// TIA Portal project "Plc_KTKDL" (V19)

(* hardware
DEVICE "S7-1200 station_1"  S7-1200 Station
   slot 0: "Rack_0"  S7-1200 Rack  Rack  V1.0
   slot 1: "PLC_1"  CPU 1214C DC/DC/DC  6ES7 214-1AG40-0XB0  V4.0
DEVICE "PC-System_1"  SIMATIC PC station
   slot 0: "SIMATIC PC station"  Rail  SIMATIC PC-Station  V1.0
      slot 125: "Stationmanager"  Station_Manager  V6.0.4
   slot 1: "HMI_RT_1"  WinCC Unified PC RT  6AV2 155-xxxxx-xxxx  19.0.0.0
   slot 2: "IE general_1"  IE General  IE_CP  V8.2.0
      slot 1: "PROFINET interface"  IEGeneral.Interface.8.2.0
*)

// ===== PLC "PLC_1"  CPU 1214C DC/DC/DC =====

VAR_GLOBAL   // PLC tag table "Default tag table"
   "Step_Lift_Pulse" AT %Q0.0 : Bool;
   "Step_Lift_Direction" AT %Q0.1 : Bool;
   "Step_Reach_Pulse" AT %Q0.4 : Bool;
   "Step_Reach_Direction" AT %Q0.5 : Bool;
   "Axis_1_Direction" AT %Q0.3 : Bool;
   "Axis_1_Pulse" AT %Q0.2 : Bool;
   "Step_Lift_Homing switch" AT %I0.0 : Bool;
END_VAR

VAR_GLOBAL   // PLC tag table "Input"
   "SensorHome" AT %M0.1 : Bool;
END_VAR

TYPE "UDT"
   STRUCT
      Monitor : Struct
         Velocity : Real;
         Position : Real;
      END_STRUCT;
      Job : Struct
         Velocity : Real;
         Forwork : Bool;
         Backwork : Bool;
         Erorr : Bool;
      END_STRUCT;
      StaticAxis : Int;
   END_STRUCT;
END_TYPE

DATA_BLOCK "DB_Vị_trí_xe"   // DB2
{ S7_Optimized_Access := 'FALSE' }
VERSION : 0.1
   VAR
      "vị trí 1" : Bool;
      "vị trí 2" : Bool;
      "vị trí 3" : Bool;
      "vị trí 4" : Bool;
      "vị trí 5" : Bool;
      "vị trí 6" : Bool;
      "vị trí 7" : Bool;
      "vị trí 8" : Bool;
      tầng_1 : Bool;
      tầng_2 : Bool;
   END_VAR
BEGIN
END_DATA_BLOCK

DATA_BLOCK "P_Trig"   // DB3
{ S7_Optimized_Access := 'TRUE' }
VERSION : 0.1
   VAR
      CLK : Array[0..100] of Bool;
   END_VAR
BEGIN
END_DATA_BLOCK

DATA_BLOCK "DB_AxisPanel"   // DB5
{ S7_Optimized_Access := 'TRUE' }
VERSION : 0.1
   VAR
      Lift : "UDT";
      Rotation : "UDT";
      Reach : "UDT";
   END_VAR
BEGIN
END_DATA_BLOCK

DATA_BLOCK "DB_Operater"   // DB6
{ S7_Optimized_Access := 'FALSE' }
VERSION : 0.1
   VAR
      Confirm_Gửi : Bool;
      Confirm_Lấy : Bool;
      ConfirmRFID : Bool;
      Scada_Gửi_Xe : Bool;
      Scada_Lấy_Xe : Bool;
      Scada_RFID : Bool;
      Scada_Home_Lift : Bool;
      BackHome : Bool;
      "Auto/Man" : Bool;
      Static_Mode : Int;
   END_VAR
BEGIN
END_DATA_BLOCK

DATA_BLOCK "DB_Convert"   // DB14
{ S7_Optimized_Access := 'FALSE' }
VERSION : 0.1
   VAR
      Python : Struct
         Floor : Int := 0;
         Location : Int;
         Passcodeplc : Int;
         UID : Array[1..12] of String[14];
         Receive : String[14];
      END_STRUCT;
      Floor_Dic1 : Int;
      Floor_Dic2 : Int;
      Location : Int;
      Down : Int;
      Up : Int;
      Started : Bool;
   END_VAR
BEGIN
END_DATA_BLOCK

// folder: Step

DATA_BLOCK "DB_Step"   // DB15
{ S7_Optimized_Access := 'TRUE' }
VERSION : 0.1
   VAR
      Power : Bool;
      Home : Struct
         Lift : Bool;
         Rotation : Bool;
         Reach : Bool;
      END_STRUCT;
      HomeAll : Bool;
      ErorrHomeCode : Struct
         Lift : Word;
         Rotation : Word;
         Reach : Word;
      END_STRUCT;
      ErrorHome : Struct
         Lift : Bool;
         Rotation : Bool;
         Reach : Bool;
      END_STRUCT;
      ErorrAbsoluteCode : Struct
         Rotation : Word;
         Lift : Word;
         Reach : Word;
      END_STRUCT;
      ErrorAbsolute : Struct
         Lift : Bool;
         Rotation : Bool;
         Reach : Bool;
      END_STRUCT;
      ErrorJog : Struct
         Lift : Word;
         Rotation : Word;
         Reach : Word;
      END_STRUCT;
      Reset : Bool;
      PowerStarted : Bool;
      HomeStarted : Bool;
      DoneHome : Bool;
   END_VAR
BEGIN
END_DATA_BLOCK

DATA_BLOCK "DB_Scrips"   // DB45
{ S7_Optimized_Access := 'FALSE' }
VERSION : 0.1
   VAR
      Dic : Int;
      "Step" : Int;
      Velocity : Struct
         Lift : Int;
         Rotation : Int;
         Reach : Int;
      END_STRUCT;
      Position : Struct
         Lift : Int;
         Rotation : Int;
         Reach : Int;
      END_STRUCT;
      Excute : Struct
         Lift : Bool;
         Rotation : Bool;
         Reach : Bool;
      END_STRUCT;
      ExcuteReady : Bool;
      Cònirm2 : Bool;
      Cònirm1 : Bool;
      Busy : Bool;
   END_VAR
BEGIN
END_DATA_BLOCK

// folder: System blocks/Program resources

DATA_BLOCK "DelayStep3"   // DB11
{ S7_Optimized_Access := 'TRUE' }
AUTHOR : Simatic
FAMILY : IEC
NAME : IEC_TMR
VERSION : 1.0
// stored: InstanceOfName IEC_TIMER
"IEC_TIMER"
BEGIN
END_DATA_BLOCK

DATA_BLOCK "Delay2s"   // DB23
{ S7_Optimized_Access := 'TRUE' }
AUTHOR : Simatic
FAMILY : IEC
NAME : IEC_TMR
VERSION : 1.0
// stored: InstanceOfName IEC_TIMER
"IEC_TIMER"
BEGIN
END_DATA_BLOCK

DATA_BLOCK "DelayStep4"   // DB47
{ S7_Optimized_Access := 'TRUE' }
AUTHOR : Simatic
FAMILY : IEC
NAME : IEC_TMR
VERSION : 1.0
// stored: InstanceOfName IEC_TIMER
"IEC_TIMER"
BEGIN
END_DATA_BLOCK

DATA_BLOCK "Delay1s5"   // DB49
{ S7_Optimized_Access := 'TRUE' }
AUTHOR : Simatic
FAMILY : IEC
NAME : IEC_TMR
VERSION : 1.0
// stored: InstanceOfName IEC_TIMER
"IEC_TIMER"
BEGIN
END_DATA_BLOCK

DATA_BLOCK "DelayyStep3"   // DB50
{ S7_Optimized_Access := 'TRUE' }
AUTHOR : Simatic
FAMILY : IEC
NAME : IEC_TMR
VERSION : 1.0
// stored: InstanceOfName IEC_TIMER
"IEC_TIMER"
BEGIN
END_DATA_BLOCK

// folder: đầy , các logic tìm

DATA_BLOCK "DB_Tìm&&Xácnhan"   // DB1
{ S7_Optimized_Access := 'TRUE' }
VERSION : 0.1
   VAR
      Call_tìm_vị_trí : Bool;
      Call_tìm_tầng : Bool;
      Xác_nhận_vị_trí : DInt;
      Xác_nhận_tầng : DInt;
   END_VAR
BEGIN
END_DATA_BLOCK

DATA_BLOCK "DB_đầy"   // DB4
{ S7_Optimized_Access := 'TRUE' }
VERSION : 0.1
   VAR
      Tầng1 : Bool;
      Tầng2 : Bool;
   END_VAR
BEGIN
END_DATA_BLOCK

// folder: (top level)

DATA_BLOCK "Step_Lift"   // DB10, Motion_DB
{ S7_Optimized_Access := 'TRUE' }
AUTHOR : SIMATIC
FAMILY : BasicMC
NAME : TO_PosAx
VERSION : 4.0
// stored: InstanceOfName TO_PositioningAxis
"TO_PositioningAxis"
BEGIN
   // Axis.DirectionOutputEnabledCU = TRUE
   // Axis.OnlinePtoModeCU = 16#0000_0002
   // Axis.SelectedChannel2EnumCU = %Q0.1
   // Axis.SelectedChannel1EnumCU = %Q0.0
   // Pulse.MinDeltaDeltaFrequencyCU = 0.004
   // Pulse.MaxDeltaDeltaFrequencyCU = 1.0E+10
   // Pulse.MinDeltaFrequencyCU = 0.005
   // Pulse.MaxDeltaFrequencyCU = 9.5E+9
   // Pulse.MinFrequencyCU = 1.0
   // Pulse.MaxFrequencyCU = 100000.0
   // Pulse.OutputSourceCU = 16#0000_0000
   // Axis.SelectPTO = 0
   // Axis.LengthUnitNormalized.Distance = 1013
END_DATA_BLOCK

DATA_BLOCK "Step_Reach"   // DB12, Motion_DB
{ S7_Optimized_Access := 'TRUE' }
AUTHOR : SIMATIC
FAMILY : BasicMC
NAME : TO_PosAx
VERSION : 4.0
// stored: InstanceOfName TO_PositioningAxis
"TO_PositioningAxis"
BEGIN
   // Axis.DirectionOutputEnabledCU = TRUE
   // Axis.OnlinePtoModeCU = 16#0000_0002
   // Axis.SelectedChannel2EnumCU = %Q0.5
   // Axis.SelectedChannel1EnumCU = %Q0.4
   // Pulse.MinDeltaDeltaFrequencyCU = 0.004
   // Pulse.MaxDeltaDeltaFrequencyCU = 1.0E+10
   // Pulse.MinDeltaFrequencyCU = 0.005
   // Pulse.MaxDeltaFrequencyCU = 9.5E+9
   // Pulse.MinFrequencyCU = 1.0
   // Pulse.MaxFrequencyCU = 30000.0
   // Pulse.OutputSourceCU = 16#0000_0000
   // Axis.SelectPTO = 1
   // Axis.OnlinePtoIndexCU = 1
   // Axis.LengthUnitNormalized.Distance = 1013
END_DATA_BLOCK

DATA_BLOCK "Step_Rotation"   // DB13, Motion_DB
{ S7_Optimized_Access := 'TRUE' }
AUTHOR : SIMATIC
FAMILY : BasicMC
NAME : TO_PosAx
VERSION : 4.0
// stored: InstanceOfName TO_PositioningAxis
"TO_PositioningAxis"
BEGIN
   // Axis.LengthUnitNormalized.Distance = 1005
   // Axis.LengthUnit.LastDistance = 1005
   // Axis.DirectionOutputEnabledCU = TRUE
   // Axis.OnlinePtoModeCU = 16#0000_0002
   // Axis.SelectedChannel2EnumCU = %Q0.3
   // Axis.SelectedChannel1EnumCU = %Q0.2
   // Pulse.MinDeltaDeltaFrequencyCU = 0.004
   // Pulse.MaxDeltaDeltaFrequencyCU = 1.0E+10
   // Pulse.MinDeltaFrequencyCU = 0.005
   // Pulse.MaxDeltaFrequencyCU = 9.5E+9
   // Pulse.MinFrequencyCU = 1.0
   // Pulse.MaxFrequencyCU = 100000.0
   // Pulse.OutputSourceCU = 16#0000_0000
   // Axis.SelectPTO = 2
   // Axis.OnlinePtoIndexCU = 2
END_DATA_BLOCK

FUNCTION "FC_SendPython" : Void   // FC1, LAD
{ S7_Optimized_Access := 'TRUE' }
VERSION : 0.1
BEGIN

REGION Network 1
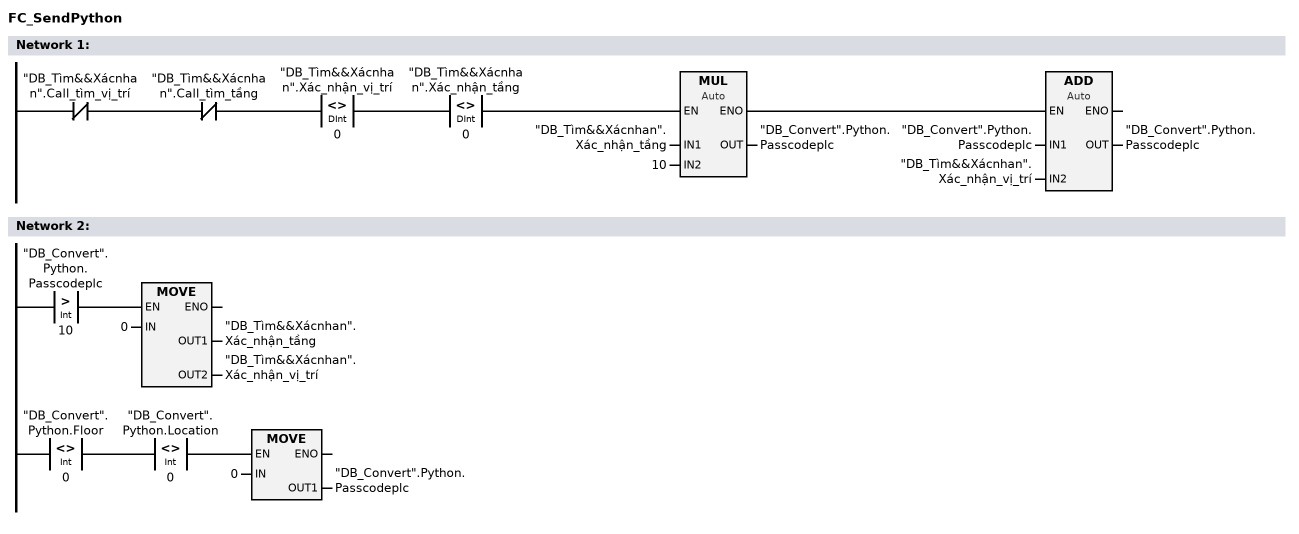
   RUNG wire#powerrail
      I_Contact( "DB_Tìm&&Xácnhan".Call_tìm_vị_trí )
      I_Contact( "DB_Tìm&&Xácnhan".Call_tìm_tầng )
      { S7_Templates := "SrcType := DInt" } NE_Contact(in1 := "DB_Tìm&&Xácnhan".Xác_nhận_vị_trí, in2 := 0)
      { S7_Templates := "SrcType := DInt" } NE_Contact(in1 := "DB_Tìm&&Xácnhan".Xác_nhận_tầng, in2 := 0)
      Mul(in1 := "DB_Tìm&&Xácnhan".Xác_nhận_tầng, in2 := 10, out => "DB_Convert".Python.Passcodeplc)
      Add(in1 := "DB_Convert".Python.Passcodeplc, in2 := "DB_Tìm&&Xácnhan".Xác_nhận_vị_trí, out => "DB_Convert".Python.Passcodeplc)
   END_RUNG
   // the same network as SCL:
   IF NOT "DB_Tìm&&Xácnhan".Call_tìm_vị_trí AND NOT "DB_Tìm&&Xácnhan".Call_tìm_tầng AND ("DB_Tìm&&Xácnhan".Xác_nhận_vị_trí <> 0) AND ("DB_Tìm&&Xácnhan".Xác_nhận_tầng <> 0) THEN
       "DB_Convert".Python.Passcodeplc := "DB_Tìm&&Xácnhan".Xác_nhận_tầng * 10;
       "DB_Convert".Python.Passcodeplc := "DB_Convert".Python.Passcodeplc + "DB_Tìm&&Xácnhan".Xác_nhận_vị_trí;
   END_IF;
END_REGION

REGION Network 2
   RUNG wire#powerrail
      { S7_Templates := "SrcType := Int" } GT_Contact(in1 := "DB_Convert".Python.Passcodeplc, in2 := 10)
      Move(in := 0, out1 => "DB_Tìm&&Xácnhan".Xác_nhận_tầng, out2 => "DB_Tìm&&Xácnhan".Xác_nhận_vị_trí)
   END_RUNG
   RUNG wire#powerrail
      { S7_Templates := "SrcType := Int" } NE_Contact(in1 := "DB_Convert".Python.Floor, in2 := 0)
      { S7_Templates := "SrcType := Int" } NE_Contact(in1 := "DB_Convert".Python.Location, in2 := 0)
      Move(in := 0, out1 => "DB_Convert".Python.Passcodeplc)
   END_RUNG
   // the same network as SCL:
   IF "DB_Convert".Python.Passcodeplc > 10 THEN
       "DB_Tìm&&Xácnhan".Xác_nhận_tầng := 0;
       "DB_Tìm&&Xácnhan".Xác_nhận_vị_trí := 0;
   END_IF;
   IF ("DB_Convert".Python.Floor <> 0) AND ("DB_Convert".Python.Location <> 0) THEN
       "DB_Convert".Python.Passcodeplc := 0;
   END_IF;
END_REGION
END_FUNCTION

FUNCTION "FC_Operater" : Void   // FC5, LAD
{ S7_Optimized_Access := 'TRUE' }
VERSION : 0.1
   VAR_TEMP   // added for the SCL form of the ladder/FBD networks
      _w1 : Bool;
      _w2 : Bool;
   END_VAR
BEGIN

REGION Network 1
   // chờ khi người dùng bấm rồi mới chạy
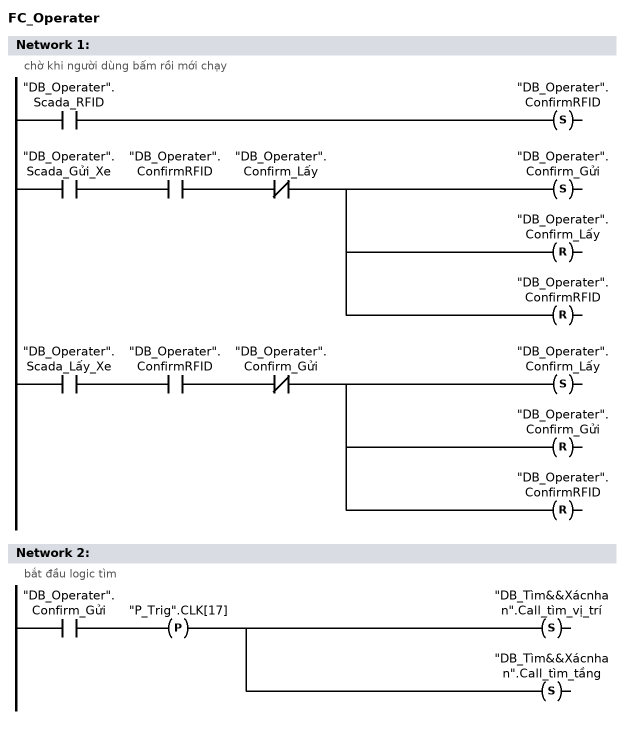
   RUNG wire#powerrail
      Contact( "DB_Operater".Scada_RFID )
      S_Coil( "DB_Operater".ConfirmRFID )
   END_RUNG
   RUNG wire#powerrail
      Contact( "DB_Operater".Scada_Gửi_Xe )
      Contact( "DB_Operater".ConfirmRFID )
      I_Contact( "DB_Operater".Confirm_Lấy )
      wire#w1
      S_Coil( "DB_Operater".Confirm_Gửi )
   END_RUNG
   RUNG wire#w1
      R_Coil( "DB_Operater".Confirm_Lấy )
   END_RUNG
   RUNG wire#w1
      R_Coil( "DB_Operater".ConfirmRFID )
   END_RUNG
   RUNG wire#powerrail
      Contact( "DB_Operater".Scada_Lấy_Xe )
      Contact( "DB_Operater".ConfirmRFID )
      I_Contact( "DB_Operater".Confirm_Gửi )
      wire#w2
      S_Coil( "DB_Operater".Confirm_Lấy )
   END_RUNG
   RUNG wire#w2
      R_Coil( "DB_Operater".Confirm_Gửi )
   END_RUNG
   RUNG wire#w2
      R_Coil( "DB_Operater".ConfirmRFID )
   END_RUNG
   // the same network as SCL:
   IF "DB_Operater".Scada_RFID THEN "DB_Operater".ConfirmRFID := TRUE; END_IF;
   IF "DB_Operater".Scada_Gửi_Xe AND "DB_Operater".ConfirmRFID AND NOT "DB_Operater".Confirm_Lấy THEN
       "DB_Operater".Confirm_Gửi := TRUE;
   END_IF;
   #_w1 := "DB_Operater".Scada_Gửi_Xe AND "DB_Operater".ConfirmRFID AND NOT "DB_Operater".Confirm_Lấy;
   IF #_w1 THEN
       "DB_Operater".Confirm_Lấy := FALSE;
       "DB_Operater".ConfirmRFID := FALSE;
   END_IF;
   IF "DB_Operater".Scada_Lấy_Xe AND "DB_Operater".ConfirmRFID AND NOT "DB_Operater".Confirm_Gửi THEN
       "DB_Operater".Confirm_Lấy := TRUE;
   END_IF;
   #_w2 := "DB_Operater".Scada_Lấy_Xe AND "DB_Operater".ConfirmRFID AND NOT "DB_Operater".Confirm_Gửi;
   IF #_w2 THEN
       "DB_Operater".Confirm_Gửi := FALSE;
       "DB_Operater".ConfirmRFID := FALSE;
   END_IF;
END_REGION

REGION Network 2
   // bắt đầu logic tìm
   RUNG wire#powerrail
      Contact( "DB_Operater".Confirm_Gửi )
      P_Trig( "P_Trig".CLK[17] )
      wire#w1
      S_Coil( "DB_Tìm&&Xácnhan".Call_tìm_vị_trí )
   END_RUNG
   RUNG wire#w1
      S_Coil( "DB_Tìm&&Xácnhan".Call_tìm_tầng )
   END_RUNG
   // the same network as SCL:
   #_w1 := "DB_Operater".Confirm_Gửi AND NOT "P_Trig".CLK[17];   // rising edge
   "P_Trig".CLK[17] := "DB_Operater".Confirm_Gửi;
   IF #_w1 THEN
       "DB_Tìm&&Xácnhan".Call_tìm_vị_trí := TRUE;
       "DB_Tìm&&Xácnhan".Call_tìm_tầng := TRUE;
   END_IF;
END_REGION
END_FUNCTION

FUNCTION "Fc_Convert" : Void   // FC7, LAD
{ S7_Optimized_Access := 'TRUE' }
VERSION : 0.1
BEGIN

REGION Network 1
   // chuyen quang duong di cua truc nang
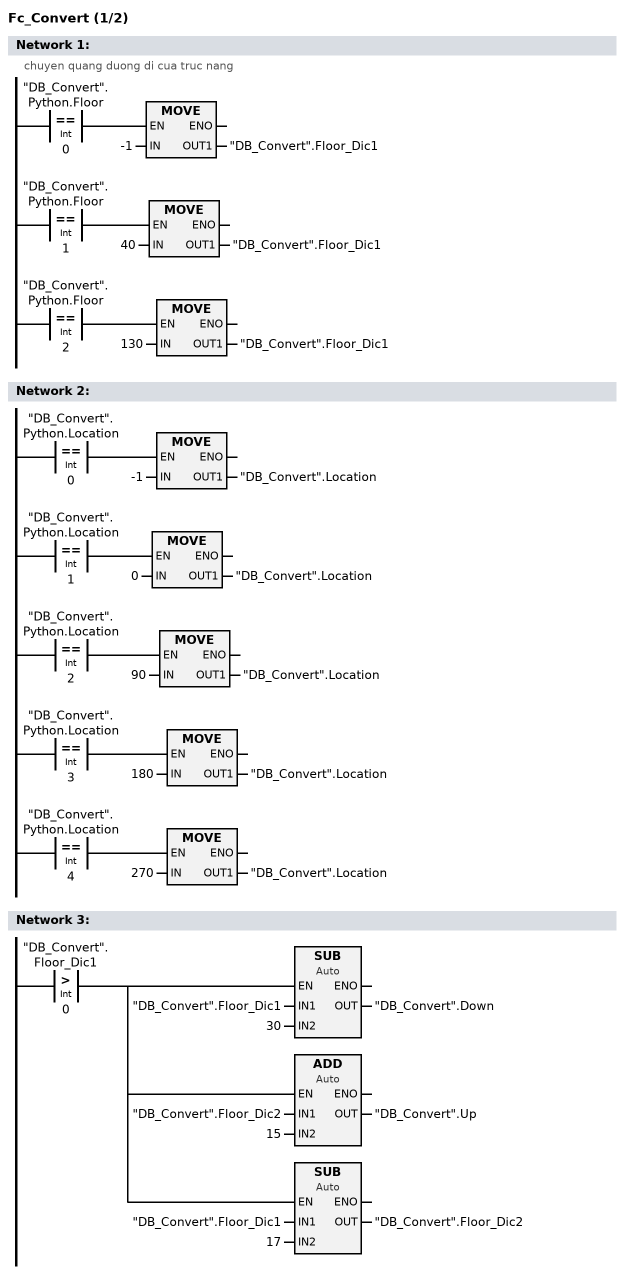
   RUNG wire#powerrail
      { S7_Templates := "SrcType := Int" } EQ_Contact(in1 := "DB_Convert".Python.Floor, in2 := 0)
      Move(in := -1, out1 => "DB_Convert".Floor_Dic1)
   END_RUNG
   RUNG wire#powerrail
      { S7_Templates := "SrcType := Int" } EQ_Contact(in1 := "DB_Convert".Python.Floor, in2 := 1)
      Move(in := 40, out1 => "DB_Convert".Floor_Dic1)
   END_RUNG
   RUNG wire#powerrail
      { S7_Templates := "SrcType := Int" } EQ_Contact(in1 := "DB_Convert".Python.Floor, in2 := 2)
      Move(in := 130, out1 => "DB_Convert".Floor_Dic1)
   END_RUNG
   // the same network as SCL:
   IF "DB_Convert".Python.Floor = 0 THEN "DB_Convert".Floor_Dic1 := -1; END_IF;
   IF "DB_Convert".Python.Floor = 1 THEN "DB_Convert".Floor_Dic1 := 40; END_IF;
   IF "DB_Convert".Python.Floor = 2 THEN "DB_Convert".Floor_Dic1 := 130; END_IF;
END_REGION

REGION Network 2
   RUNG wire#powerrail
      { S7_Templates := "SrcType := Int" } EQ_Contact(in1 := "DB_Convert".Python.Location, in2 := 0)
      Move(in := -1, out1 => "DB_Convert".Location)
   END_RUNG
   RUNG wire#powerrail
      { S7_Templates := "SrcType := Int" } EQ_Contact(in1 := "DB_Convert".Python.Location, in2 := 1)
      Move(in := 0, out1 => "DB_Convert".Location)
   END_RUNG
   RUNG wire#powerrail
      { S7_Templates := "SrcType := Int" } EQ_Contact(in1 := "DB_Convert".Python.Location, in2 := 2)
      Move(in := 90, out1 => "DB_Convert".Location)
   END_RUNG
   RUNG wire#powerrail
      { S7_Templates := "SrcType := Int" } EQ_Contact(in1 := "DB_Convert".Python.Location, in2 := 3)
      Move(in := 180, out1 => "DB_Convert".Location)
   END_RUNG
   RUNG wire#powerrail
      { S7_Templates := "SrcType := Int" } EQ_Contact(in1 := "DB_Convert".Python.Location, in2 := 4)
      Move(in := 270, out1 => "DB_Convert".Location)
   END_RUNG
   // the same network as SCL:
   IF "DB_Convert".Python.Location = 0 THEN "DB_Convert".Location := -1; END_IF;
   IF "DB_Convert".Python.Location = 1 THEN "DB_Convert".Location := 0; END_IF;
   IF "DB_Convert".Python.Location = 2 THEN "DB_Convert".Location := 90; END_IF;
   IF "DB_Convert".Python.Location = 3 THEN "DB_Convert".Location := 180; END_IF;
   IF "DB_Convert".Python.Location = 4 THEN "DB_Convert".Location := 270; END_IF;
END_REGION

REGION Network 3
   RUNG wire#powerrail
      { S7_Templates := "SrcType := Int" } GT_Contact(in1 := "DB_Convert".Floor_Dic1, in2 := 0)
      wire#w1
      Sub(in1 := "DB_Convert".Floor_Dic1, in2 := 30, out => "DB_Convert".Down)
   END_RUNG
   RUNG wire#w1
      Add(in1 := "DB_Convert".Floor_Dic2, in2 := 15, out => "DB_Convert".Up)
   END_RUNG
   RUNG wire#w1
      Sub(in1 := "DB_Convert".Floor_Dic1, in2 := 17, out => "DB_Convert".Floor_Dic2)
   END_RUNG
   // the same network as SCL:
   IF "DB_Convert".Floor_Dic1 > 0 THEN
       "DB_Convert".Down := "DB_Convert".Floor_Dic1 - 30;
       "DB_Convert".Up := "DB_Convert".Floor_Dic2 + 15;
       "DB_Convert".Floor_Dic2 := "DB_Convert".Floor_Dic1 - 17;
   END_IF;
END_REGION

REGION Network 4
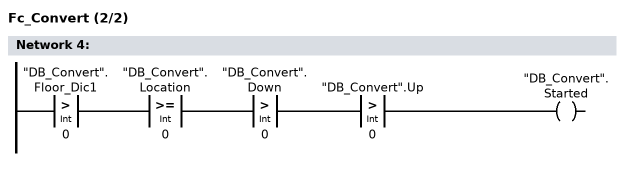
   RUNG wire#powerrail
      { S7_Templates := "SrcType := Int" } GT_Contact(in1 := "DB_Convert".Floor_Dic1, in2 := 0)
      { S7_Templates := "SrcType := Int" } GE_Contact(in1 := "DB_Convert".Location, in2 := 0)
      { S7_Templates := "SrcType := Int" } GT_Contact(in1 := "DB_Convert".Down, in2 := 0)
      { S7_Templates := "SrcType := Int" } GT_Contact(in1 := "DB_Convert".Up, in2 := 0)
      Coil( "DB_Convert".Started )
   END_RUNG
   // the same network as SCL:
   "DB_Convert".Started := ("DB_Convert".Floor_Dic1 > 0) AND ("DB_Convert".Location >= 0) AND ("DB_Convert".Down > 0) AND ("DB_Convert".Up > 0);
END_REGION
END_FUNCTION

FUNCTION "FC_Manual" : Void   // FC9, LAD
{ S7_Optimized_Access := 'TRUE' }
VERSION : 0.1
   VAR_TEMP   // added for the SCL form of the ladder/FBD networks
      _w1 : Bool;
   END_VAR
BEGIN

REGION Network 1
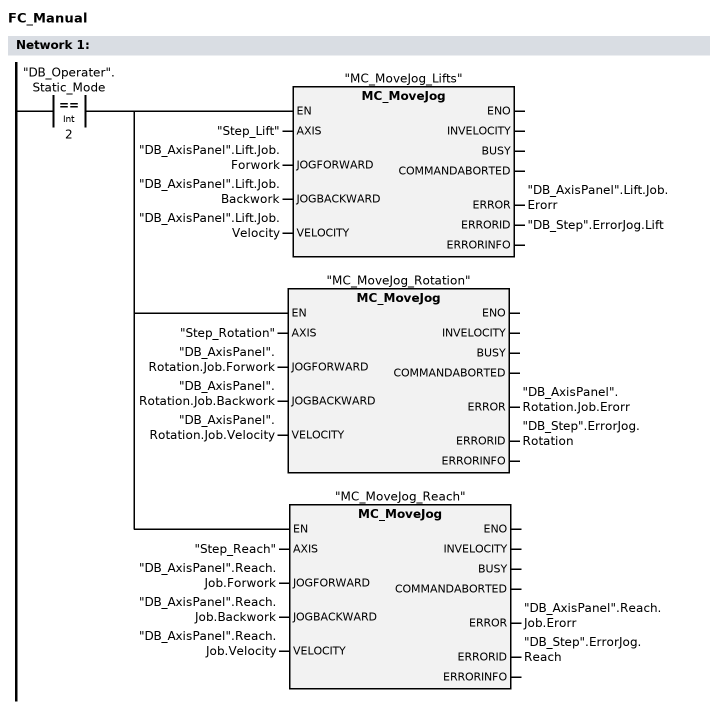
   #_w1 := "DB_Operater".Static_Mode = 2;
   IF #_w1 THEN
       "MC_MoveJog_Lifts"(Axis := "Step_Lift",   // MC_MoveJog
                          JogForward := "DB_AxisPanel".Lift.Job.Forwork,
                          JogBackward := "DB_AxisPanel".Lift.Job.Backwork,
                          Velocity := "DB_AxisPanel".Lift.Job.Velocity,
                          Error => "DB_AxisPanel".Lift.Job.Erorr,
                          ErrorID => "DB_Step".ErrorJog.Lift);
       "MC_MoveJog_Rotation"(Axis := "Step_Rotation",   // MC_MoveJog
                             JogForward := "DB_AxisPanel".Rotation.Job.Forwork,
                             JogBackward := "DB_AxisPanel".Rotation.Job.Backwork,
                             Velocity := "DB_AxisPanel".Rotation.Job.Velocity,
                             Error => "DB_AxisPanel".Rotation.Job.Erorr,
                             ErrorID => "DB_Step".ErrorJog.Rotation);
       "MC_MoveJog_Reach"(Axis := "Step_Reach",   // MC_MoveJog
                          JogForward := "DB_AxisPanel".Reach.Job.Forwork,
                          JogBackward := "DB_AxisPanel".Reach.Job.Backwork,
                          Velocity := "DB_AxisPanel".Reach.Job.Velocity,
                          Error => "DB_AxisPanel".Reach.Job.Erorr,
                          ErrorID => "DB_Step".ErrorJog.Reach);
   END_IF;
END_REGION
END_FUNCTION

FUNCTION "FC_PanelAxis" : Void   // FC10, LAD
{ S7_Optimized_Access := 'TRUE' }
VERSION : 0.1
BEGIN

REGION Network 1
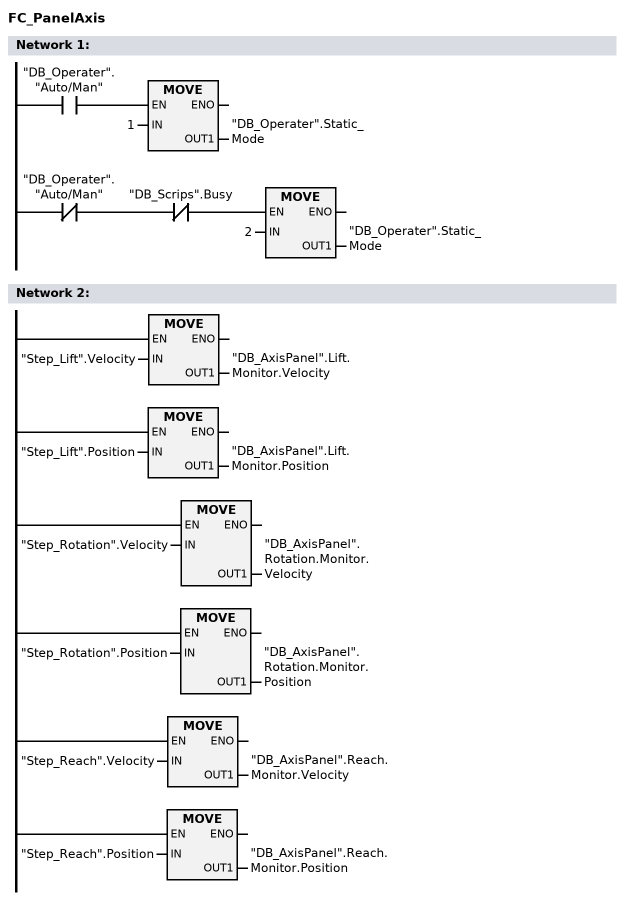
   RUNG wire#powerrail
      Contact( "DB_Operater"."Auto/Man" )
      Move(in := 1, out1 => "DB_Operater".Static_Mode)
   END_RUNG
   RUNG wire#powerrail
      I_Contact( "DB_Operater"."Auto/Man" )
      I_Contact( "DB_Scrips".Busy )
      Move(in := 2, out1 => "DB_Operater".Static_Mode)
   END_RUNG
   // the same network as SCL:
   IF "DB_Operater"."Auto/Man" THEN "DB_Operater".Static_Mode := 1; END_IF;
   IF NOT "DB_Operater"."Auto/Man" AND NOT "DB_Scrips".Busy THEN "DB_Operater".Static_Mode := 2; END_IF;
END_REGION

REGION Network 2
   RUNG wire#powerrail
      Move(in := "Step_Lift".Velocity, out1 => "DB_AxisPanel".Lift.Monitor.Velocity)
   END_RUNG
   RUNG wire#powerrail
      Move(in := "Step_Lift".Position, out1 => "DB_AxisPanel".Lift.Monitor.Position)
   END_RUNG
   RUNG wire#powerrail
      Move(in := "Step_Rotation".Velocity, out1 => "DB_AxisPanel".Rotation.Monitor.Velocity)
   END_RUNG
   RUNG wire#powerrail
      Move(in := "Step_Rotation".Position, out1 => "DB_AxisPanel".Rotation.Monitor.Position)
   END_RUNG
   RUNG wire#powerrail
      Move(in := "Step_Reach".Velocity, out1 => "DB_AxisPanel".Reach.Monitor.Velocity)
   END_RUNG
   RUNG wire#powerrail
      Move(in := "Step_Reach".Position, out1 => "DB_AxisPanel".Reach.Monitor.Position)
   END_RUNG
   // the same network as SCL:
   "DB_AxisPanel".Lift.Monitor.Velocity := "Step_Lift".Velocity;
   "DB_AxisPanel".Lift.Monitor.Position := "Step_Lift".Position;
   "DB_AxisPanel".Rotation.Monitor.Velocity := "Step_Rotation".Velocity;
   "DB_AxisPanel".Rotation.Monitor.Position := "Step_Rotation".Position;
   "DB_AxisPanel".Reach.Monitor.Velocity := "Step_Reach".Velocity;
   "DB_AxisPanel".Reach.Monitor.Position := "Step_Reach".Position;
END_REGION
END_FUNCTION

FUNCTION "FC_BackHome" : Void   // FC11, LAD
{ S7_Optimized_Access := 'TRUE' }
VERSION : 0.1
BEGIN
END_FUNCTION

FUNCTION "FC_UID" : Void   // FC12, LAD
{ S7_Optimized_Access := 'TRUE' }
VERSION : 0.1
   VAR_TEMP   // added for the SCL form of the ladder/FBD networks
      _w1 : Bool;
      _w2 : Bool;
      _w3 : Bool;
   END_VAR
BEGIN

REGION Network 1
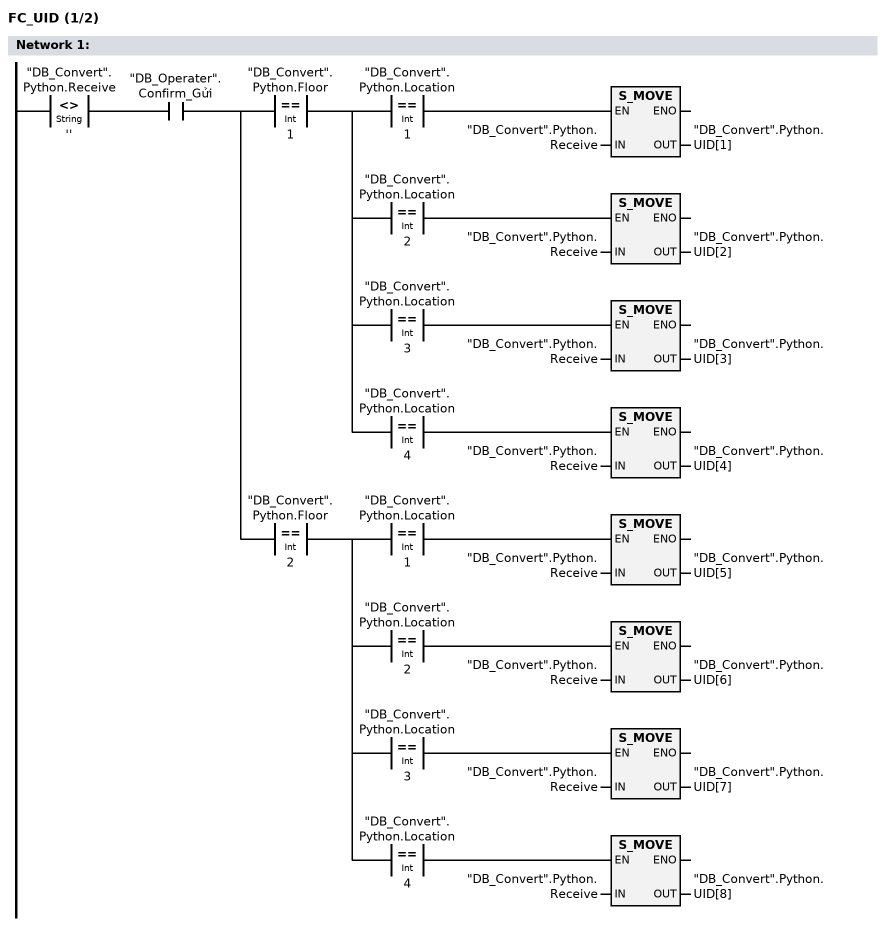
   RUNG wire#powerrail
      { S7_Templates := "SrcType := String" } NE_Contact(in1 := "DB_Convert".Python.Receive, in2 := '')
      Contact( "DB_Operater".Confirm_Gửi )
      wire#w1
      { S7_Templates := "SrcType := Int" } EQ_Contact(in1 := "DB_Convert".Python.Floor, in2 := 1)
      wire#w2
      { S7_Templates := "SrcType := Int" } EQ_Contact(in1 := "DB_Convert".Python.Location, in2 := 1)
      S_Move(in := "DB_Convert".Python.Receive, out => "DB_Convert".Python.UID[1])
   END_RUNG
   RUNG wire#w2
      { S7_Templates := "SrcType := Int" } EQ_Contact(in1 := "DB_Convert".Python.Location, in2 := 2)
      S_Move(in := "DB_Convert".Python.Receive, out => "DB_Convert".Python.UID[2])
   END_RUNG
   RUNG wire#w2
      { S7_Templates := "SrcType := Int" } EQ_Contact(in1 := "DB_Convert".Python.Location, in2 := 3)
      S_Move(in := "DB_Convert".Python.Receive, out => "DB_Convert".Python.UID[3])
   END_RUNG
   RUNG wire#w2
      { S7_Templates := "SrcType := Int" } EQ_Contact(in1 := "DB_Convert".Python.Location, in2 := 4)
      S_Move(in := "DB_Convert".Python.Receive, out => "DB_Convert".Python.UID[4])
   END_RUNG
   RUNG wire#w1
      { S7_Templates := "SrcType := Int" } EQ_Contact(in1 := "DB_Convert".Python.Floor, in2 := 2)
      wire#w3
      { S7_Templates := "SrcType := Int" } EQ_Contact(in1 := "DB_Convert".Python.Location, in2 := 1)
      S_Move(in := "DB_Convert".Python.Receive, out => "DB_Convert".Python.UID[5])
   END_RUNG
   RUNG wire#w3
      { S7_Templates := "SrcType := Int" } EQ_Contact(in1 := "DB_Convert".Python.Location, in2 := 2)
      S_Move(in := "DB_Convert".Python.Receive, out => "DB_Convert".Python.UID[6])
   END_RUNG
   RUNG wire#w3
      { S7_Templates := "SrcType := Int" } EQ_Contact(in1 := "DB_Convert".Python.Location, in2 := 3)
      S_Move(in := "DB_Convert".Python.Receive, out => "DB_Convert".Python.UID[7])
   END_RUNG
   RUNG wire#w3
      { S7_Templates := "SrcType := Int" } EQ_Contact(in1 := "DB_Convert".Python.Location, in2 := 4)
      S_Move(in := "DB_Convert".Python.Receive, out => "DB_Convert".Python.UID[8])
   END_RUNG
   // the same network as SCL:
   #_w1 := ("DB_Convert".Python.Receive <> '') AND "DB_Operater".Confirm_Gửi;
   #_w2 := #_w1 AND ("DB_Convert".Python.Floor = 1);
   IF #_w2 AND ("DB_Convert".Python.Location = 1) THEN
       "DB_Convert".Python.UID[1] := "DB_Convert".Python.Receive;
   END_IF;
   IF #_w2 AND ("DB_Convert".Python.Location = 2) THEN
       "DB_Convert".Python.UID[2] := "DB_Convert".Python.Receive;
   END_IF;
   IF #_w2 AND ("DB_Convert".Python.Location = 3) THEN
       "DB_Convert".Python.UID[3] := "DB_Convert".Python.Receive;
   END_IF;
   IF #_w2 AND ("DB_Convert".Python.Location = 4) THEN
       "DB_Convert".Python.UID[4] := "DB_Convert".Python.Receive;
   END_IF;
   #_w3 := #_w1 AND ("DB_Convert".Python.Floor = 2);
   IF #_w3 AND ("DB_Convert".Python.Location = 1) THEN
       "DB_Convert".Python.UID[5] := "DB_Convert".Python.Receive;
   END_IF;
   IF #_w3 AND ("DB_Convert".Python.Location = 2) THEN
       "DB_Convert".Python.UID[6] := "DB_Convert".Python.Receive;
   END_IF;
   IF #_w3 AND ("DB_Convert".Python.Location = 3) THEN
       "DB_Convert".Python.UID[7] := "DB_Convert".Python.Receive;
   END_IF;
   IF #_w3 AND ("DB_Convert".Python.Location = 4) THEN
       "DB_Convert".Python.UID[8] := "DB_Convert".Python.Receive;
   END_IF;
END_REGION

REGION Network 2
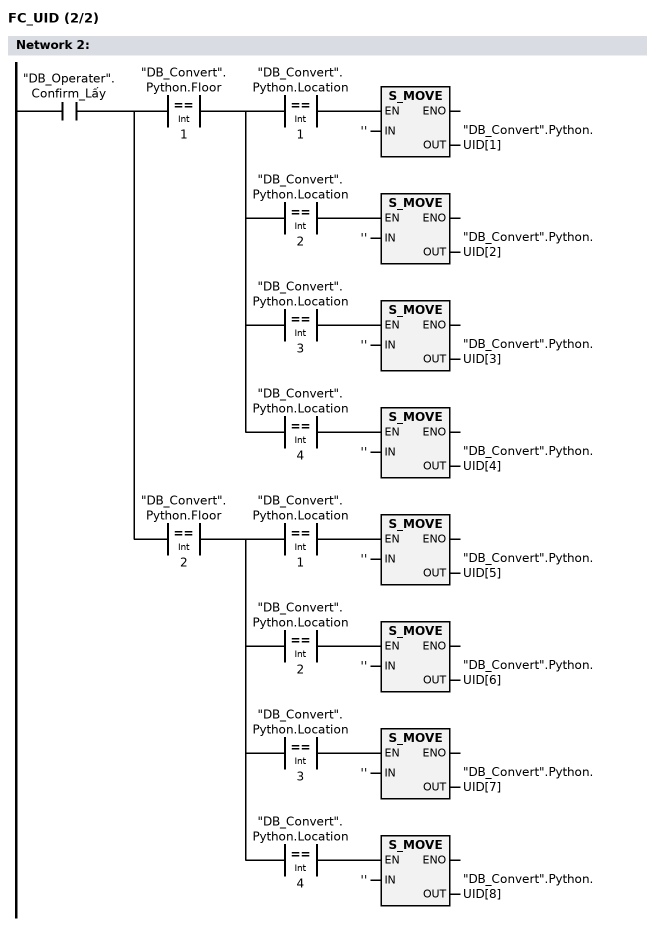
   RUNG wire#powerrail
      Contact( "DB_Operater".Confirm_Lấy )
      wire#w1
      { S7_Templates := "SrcType := Int" } EQ_Contact(in1 := "DB_Convert".Python.Floor, in2 := 1)
      wire#w2
      { S7_Templates := "SrcType := Int" } EQ_Contact(in1 := "DB_Convert".Python.Location, in2 := 1)
      S_Move(in := '', out => "DB_Convert".Python.UID[1])
   END_RUNG
   RUNG wire#w2
      { S7_Templates := "SrcType := Int" } EQ_Contact(in1 := "DB_Convert".Python.Location, in2 := 2)
      S_Move(in := '', out => "DB_Convert".Python.UID[2])
   END_RUNG
   RUNG wire#w2
      { S7_Templates := "SrcType := Int" } EQ_Contact(in1 := "DB_Convert".Python.Location, in2 := 3)
      S_Move(in := '', out => "DB_Convert".Python.UID[3])
   END_RUNG
   RUNG wire#w2
      { S7_Templates := "SrcType := Int" } EQ_Contact(in1 := "DB_Convert".Python.Location, in2 := 4)
      S_Move(in := '', out => "DB_Convert".Python.UID[4])
   END_RUNG
   RUNG wire#w1
      { S7_Templates := "SrcType := Int" } EQ_Contact(in1 := "DB_Convert".Python.Floor, in2 := 2)
      wire#w3
      { S7_Templates := "SrcType := Int" } EQ_Contact(in1 := "DB_Convert".Python.Location, in2 := 1)
      S_Move(in := '', out => "DB_Convert".Python.UID[5])
   END_RUNG
   RUNG wire#w3
      { S7_Templates := "SrcType := Int" } EQ_Contact(in1 := "DB_Convert".Python.Location, in2 := 2)
      S_Move(in := '', out => "DB_Convert".Python.UID[6])
   END_RUNG
   RUNG wire#w3
      { S7_Templates := "SrcType := Int" } EQ_Contact(in1 := "DB_Convert".Python.Location, in2 := 3)
      S_Move(in := '', out => "DB_Convert".Python.UID[7])
   END_RUNG
   RUNG wire#w3
      { S7_Templates := "SrcType := Int" } EQ_Contact(in1 := "DB_Convert".Python.Location, in2 := 4)
      S_Move(in := '', out => "DB_Convert".Python.UID[8])
   END_RUNG
   // the same network as SCL:
   #_w1 := "DB_Operater".Confirm_Lấy AND ("DB_Convert".Python.Floor = 1);
   IF #_w1 AND ("DB_Convert".Python.Location = 1) THEN "DB_Convert".Python.UID[1] := ''; END_IF;
   IF #_w1 AND ("DB_Convert".Python.Location = 2) THEN "DB_Convert".Python.UID[2] := ''; END_IF;
   IF #_w1 AND ("DB_Convert".Python.Location = 3) THEN "DB_Convert".Python.UID[3] := ''; END_IF;
   IF #_w1 AND ("DB_Convert".Python.Location = 4) THEN "DB_Convert".Python.UID[4] := ''; END_IF;
   #_w2 := "DB_Operater".Confirm_Lấy AND ("DB_Convert".Python.Floor = 2);
   IF #_w2 AND ("DB_Convert".Python.Location = 1) THEN "DB_Convert".Python.UID[5] := ''; END_IF;
   IF #_w2 AND ("DB_Convert".Python.Location = 2) THEN "DB_Convert".Python.UID[6] := ''; END_IF;
   IF #_w2 AND ("DB_Convert".Python.Location = 3) THEN "DB_Convert".Python.UID[7] := ''; END_IF;
   IF #_w2 AND ("DB_Convert".Python.Location = 4) THEN "DB_Convert".Python.UID[8] := ''; END_IF;
END_REGION
END_FUNCTION

FUNCTION "FC_Step" : Void   // FC13, LAD
{ S7_Optimized_Access := 'TRUE' }
VERSION : 0.1
   VAR_TEMP   // added for the SCL form of the ladder/FBD networks
      _w1 : Bool;
   END_VAR
BEGIN

REGION Network 1
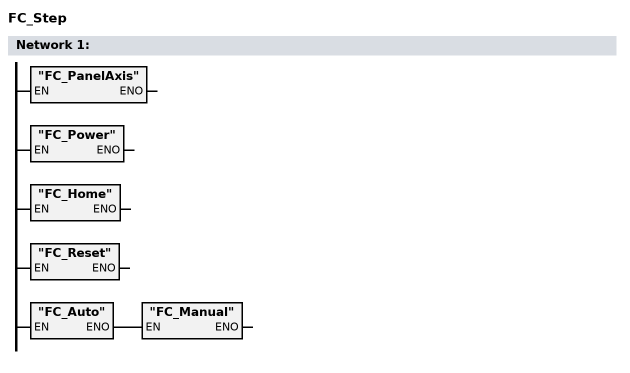
   RUNG wire#powerrail
      "FC_PanelAxis"()
   END_RUNG
   RUNG wire#powerrail
      "FC_Power"()
   END_RUNG
   RUNG wire#powerrail
      "FC_Home"()
   END_RUNG
   RUNG wire#powerrail
      "FC_Reset"()
   END_RUNG
   RUNG wire#powerrail
      "FC_Auto"()
      "FC_Manual"()
   END_RUNG
   // the same network as SCL:
   "FC_PanelAxis"();
   "FC_Power"();
   "FC_Home"();
   "FC_Reset"();
   "FC_Auto"(ENO => #_w1);
   IF #_w1 THEN "FC_Manual"(); END_IF;
END_REGION

REGION Network 2
   // Move Job
END_REGION
END_FUNCTION

FUNCTION "FC_Find" : Void   // FC14, LAD
{ S7_Optimized_Access := 'TRUE' }
VERSION : 0.1
BEGIN

REGION Network 1
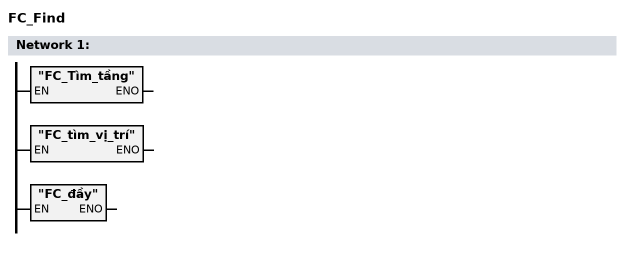
   RUNG wire#powerrail
      "FC_Tìm_tầng"()
   END_RUNG
   RUNG wire#powerrail
      "FC_tìm_vị_trí"()
   END_RUNG
   RUNG wire#powerrail
      "FC_đầy"()
   END_RUNG
   // the same network as SCL:
   "FC_Tìm_tầng"();
   "FC_tìm_vị_trí"();
   "FC_đầy"();
END_REGION
END_FUNCTION

ORGANIZATION_BLOCK "Main"   // OB1, LAD, ProgramCycle
TITLE = "Main Program Sweep (Cycle)"
{ S7_Optimized_Access := 'TRUE' }
VERSION : 0.1
   VAR_INPUT
      Initial_Call : Bool;   // Initial call of this OB
      Remanence : Bool;   // =True, if remanent data are available
   END_VAR
BEGIN

REGION Network 1
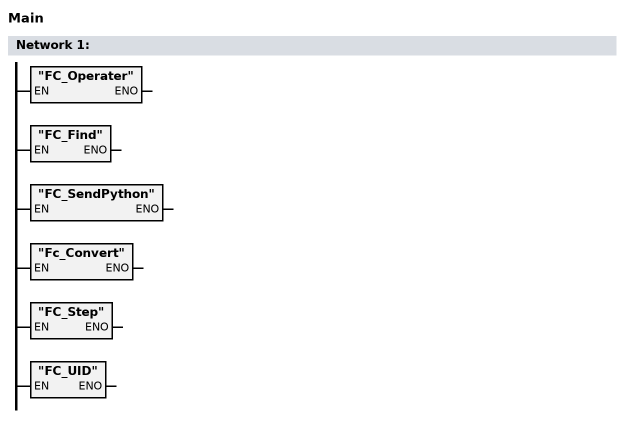
   RUNG wire#powerrail
      "FC_Operater"()
   END_RUNG
   RUNG wire#powerrail
      "FC_Find"()
   END_RUNG
   RUNG wire#powerrail
      "FC_SendPython"()
   END_RUNG
   RUNG wire#powerrail
      "Fc_Convert"()
   END_RUNG
   RUNG wire#powerrail
      "FC_Step"()
   END_RUNG
   RUNG wire#powerrail
      "FC_UID"()
   END_RUNG
   // the same network as SCL:
   "FC_Operater"();
   "FC_Find"();
   "FC_SendPython"();
   "Fc_Convert"();
   "FC_Step"();
   "FC_UID"();
END_REGION
END_ORGANIZATION_BLOCK

// folder: Step

FUNCTION "FC_Power" : Void   // FC15, LAD
{ S7_Optimized_Access := 'TRUE' }
VERSION : 0.1
BEGIN

REGION Network 1
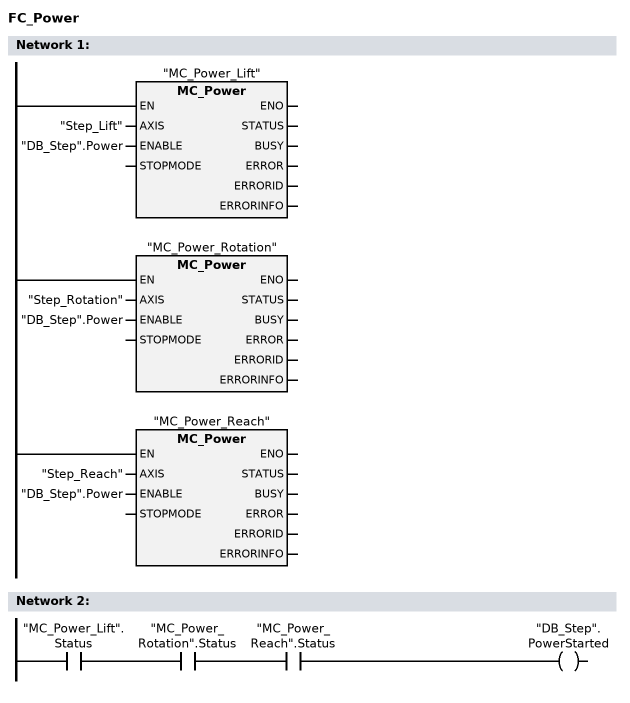
   "MC_Power_Lift"(Axis := "Step_Lift", Enable := "DB_Step".Power);   // MC_Power
   "MC_Power_Rotation"(Axis := "Step_Rotation", Enable := "DB_Step".Power);   // MC_Power
   "MC_Power_Reach"(Axis := "Step_Reach", Enable := "DB_Step".Power);   // MC_Power
END_REGION

REGION Network 2
   RUNG wire#powerrail
      Contact( "MC_Power_Lift".Status )
      Contact( "MC_Power_Rotation".Status )
      Contact( "MC_Power_Reach".Status )
      Coil( "DB_Step".PowerStarted )
   END_RUNG
   // the same network as SCL:
   "DB_Step".PowerStarted := "MC_Power_Lift".Status AND "MC_Power_Rotation".Status AND "MC_Power_Reach".Status;
END_REGION
END_FUNCTION

FUNCTION "FC_Home" : Void   // FC16, LAD
{ S7_Optimized_Access := 'TRUE' }
VERSION : 0.1
BEGIN

REGION Network 1